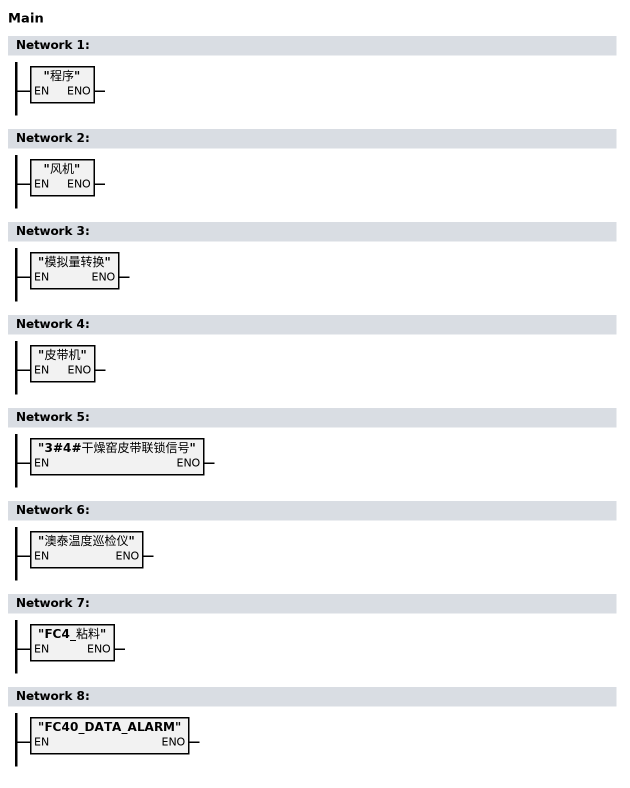
   RUNG wire#powerrail
      "程序"()
   END_RUNG
   // the same network as SCL:
   "程序"();
END_REGION

REGION Network 2
   RUNG wire#powerrail
      "风机"()
   END_RUNG
   // the same network as SCL:
   "风机"();
END_REGION

REGION Network 3
   RUNG wire#powerrail
      "模拟量转换"()
   END_RUNG
   // the same network as SCL:
   "模拟量转换"();
END_REGION

REGION Network 4
   RUNG wire#powerrail
      "皮带机"()
   END_RUNG
   // the same network as SCL:
   "皮带机"();
END_REGION

REGION Network 5
   RUNG wire#powerrail
      "3#4#干燥窑皮带联锁信号"()
   END_RUNG
   // the same network as SCL:
   "3#4#干燥窑皮带联锁信号"();
END_REGION

REGION Network 6
   RUNG wire#powerrail
      "澳泰温度巡检仪"()
   END_RUNG
   // the same network as SCL:
   "澳泰温度巡检仪"();
END_REGION

REGION Network 7
   RUNG wire#powerrail
      "FC4_粘料"()
   END_RUNG
   // the same network as SCL:
   "FC4_粘料"();
END_REGION

REGION Network 8
   RUNG wire#powerrail
      "FC40_DATA_ALARM"()
   END_RUNG
   // the same network as SCL:
   "FC40_DATA_ALARM"();
END_REGION
END_ORGANIZATION_BLOCK

ORGANIZATION_BLOCK "Cyclic interrupt"   // OB30, LAD, CyclicInterrupt
{ S7_Optimized_Access := 'TRUE' }
VERSION : 0.1
   VAR_INPUT
      Initial_Call : Bool;   // Initial call of this OB
      Event_Count : Int;   // Events discarded
   END_VAR
   VAR_TEMP   // added for the SCL form of the ladder/FBD networks
      _w1 : Bool;
      _w2 : Bool;
   END_VAR
BEGIN

REGION Network 1
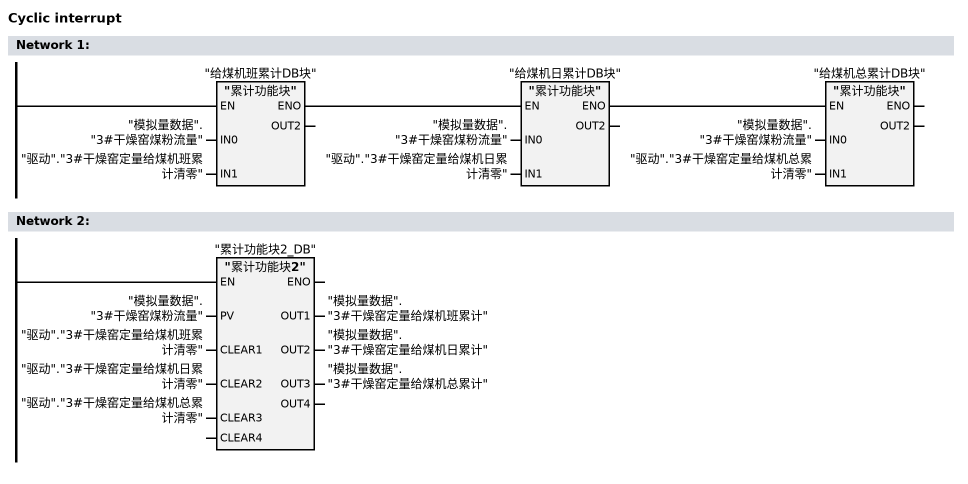
   RUNG wire#powerrail
      "给煤机班累计DB块"(IN0 := "模拟量数据"."3#干燥窑煤粉流量", IN1 := "驱动"."3#干燥窑定量给煤机班累计清零", OUT2 =>)
      "给煤机日累计DB块"(IN0 := "模拟量数据"."3#干燥窑煤粉流量", IN1 := "驱动"."3#干燥窑定量给煤机日累计清零", OUT2 =>)
      "给煤机总累计DB块"(IN0 := "模拟量数据"."3#干燥窑煤粉流量", IN1 := "驱动"."3#干燥窑定量给煤机总累计清零", OUT2 =>)
   END_RUNG
   // the same network as SCL:
   "给煤机班累计DB块"(IN0 := "模拟量数据"."3#干燥窑煤粉流量", IN1 := "驱动"."3#干燥窑定量给煤机班累计清零", ENO => #_w1);   // "累计功能块"
   "给煤机日累计DB块"(EN := #_w1, IN0 := "模拟量数据"."3#干燥窑煤粉流量", IN1 := "驱动"."3#干燥窑定量给煤机日累计清零", ENO => #_w2);   // "累计功能块"
   IF #_w2 THEN
       "给煤机总累计DB块"(IN0 := "模拟量数据"."3#干燥窑煤粉流量", IN1 := "驱动"."3#干燥窑定量给煤机总累计清零");   // "累计功能块"
   END_IF;
END_REGION

REGION Network 2
   RUNG wire#powerrail
      "累计功能块2_DB"(PV := "模拟量数据"."3#干燥窑煤粉流量", CLEAR1 := "驱动"."3#干燥窑定量给煤机班累计清零", CLEAR2 := "驱动"."3#干燥窑定量给煤机日累计清零", CLEAR3 := "驱动"."3#干燥窑定量给煤机总累计清零", CLEAR4 :=, OUT1 => "模拟量数据"."3#干燥窑定量给煤机班累计", OUT2 => "模拟量数据"."3#干燥窑定量给煤机日累计", OUT3 => "模拟量数据"."3#干燥窑定量给煤机总累计", OUT4 =>)
   END_RUNG
   // the same network as SCL:
   "累计功能块2_DB"(PV := "模拟量数据"."3#干燥窑煤粉流量",   // "累计功能块2"
               CLEAR1 := "驱动"."3#干燥窑定量给煤机班累计清零",
               CLEAR2 := "驱动"."3#干燥窑定量给煤机日累计清零",
               CLEAR3 := "驱动"."3#干燥窑定量给煤机总累计清零",
               OUT1 => "模拟量数据"."3#干燥窑定量给煤机班累计",
               OUT2 => "模拟量数据"."3#干燥窑定量给煤机日累计",
               OUT3 => "模拟量数据"."3#干燥窑定量给煤机总累计");
END_REGION
END_ORGANIZATION_BLOCK

// ===== PLC "3#HZY"  CPU 1511-1 PN =====

VAR_GLOBAL   // PLC tag table "默认变量表"
   "3#回转窑启动备妥" AT %I0.0 : Bool;
   "3#回转窑主机备妥" AT %I0.1 : Bool;
   "3#回转窑主机运行" AT %I0.2 : Bool;
   "3#回转窑主机故障" AT %I0.3 : Bool;
   "3#回转窑主机合闸" AT %I0.4 : Bool;
   "3#回转窑从机备妥" AT %I0.5 : Bool;
   "3#回转窑从机运行" AT %I0.6 : Bool;
   "3#回转窑从机故障" AT %I0.7 : Bool;
   "3#回转窑从机合闸" AT %I1.0 : Bool;
   "I1_3" AT %I1.3 : Bool;
   "I1_4" AT %I1.4 : Bool;
   "I1_5" AT %I1.5 : Bool;
   "I1_6" AT %I1.6 : Bool;
   "I1_7" AT %I1.7 : Bool;
   "主机稀油中控" AT %I2.0 : Bool;
   "主机稀油1#泵运行" AT %I2.1 : Bool;
   "主机稀油2#泵运行" AT %I2.2 : Bool;
   "主机稀油油差下限" AT %I2.3 : Bool;
   "主机稀油油位上限" AT %I2.4 : Bool;
   "主机稀油油位下限" AT %I2.5 : Bool;
   "主机稀油重故障" AT %I2.6 : Bool;
   "主机稀油轻故障" AT %I2.7 : Bool;
   "从机稀油中控" AT %I3.0 : Bool;
   "从机稀油1#泵运行" AT %I3.1 : Bool;
   "从机稀油2#泵运行" AT %I3.2 : Bool;
   "从机稀油油差下限" AT %I3.3 : Bool;
   "从机稀油油位上限" AT %I3.4 : Bool;
   "从机稀油油位下限" AT %I3.5 : Bool;
   "从机稀油重故障" AT %I3.6 : Bool;
   "从机稀油轻故障" AT %I3.7 : Bool;
   "1#挡轮备妥" AT %I4.0 : Bool;
   "1#挡轮1#泵运行" AT %I4.1 : Bool;
   "1#挡轮2#泵运行" AT %I4.2 : Bool;
   "1#挡轮溢流阀运行" AT %I4.3 : Bool;
   "挡轮重故障" AT %I4.4 : Bool;
   "挡轮轻故障" AT %I4.5 : Bool;
   "窑体行程上限" AT %I5.0 : Bool;
   "窑体行程上上限" AT %I5.1 : Bool;
   "窑体行程下限" AT %I5.2 : Bool;
   "窑体行程下下限" AT %I5.3 : Bool;
   "干矿提升皮带中控" AT %I6.0 : Bool;
   "干矿提升皮带运行" AT %I6.1 : Bool;
   "干矿提升皮带故障" AT %I6.2 : Bool;
   "干矿进料皮带中控" AT %I6.3 : Bool;
   "干矿进料皮带运行" AT %I6.4 : Bool;
   "干矿进料皮带故障" AT %I6.5 : Bool;
   "尾排风机高压远程" AT %I7.0 : Bool;
   "尾排风机高压合闸" AT %I7.1 : Bool;
   "尾排风机高压分闸" AT %I7.2 : Bool;
   "尾排风机变频远程" AT %I7.4 : Bool;
   "尾排风机变频运行" AT %I7.5 : Bool;
   "尾排风机变频故障" AT %I7.6 : Bool;
   "尾排风机变频待机" AT %I7.7 : Bool;
   "转子秤中控" AT %I8.0 : Bool;
   "转子秤运行" AT %I8.1 : Bool;
   "转子秤故障" AT %I8.2 : Bool;
   "煤粉仓收尘风机中控" AT %I8.4 : Bool;
   "煤粉仓收尘风机运行" AT %I8.5 : Bool;
   "煤粉仓收尘风机故障" AT %I8.6 : Bool;
   "回转窑一次风机中控" AT %I9.0 : Bool;
   "回转窑一次风机运行" AT %I9.1 : Bool;
   "回转窑一次风机故障" AT %I9.2 : Bool;
   "回转窑二次风机中控" AT %I9.3 : Bool;
   "回转窑二次风机运行" AT %I9.4 : Bool;
   "回转窑二次风机故障" AT %I9.5 : Bool;
   "回转窑备用一次风机中控" AT %I10.0 : Bool;
   "回转窑备用一次风机运行" AT %I10.1 : Bool;
   "回转窑备用一次风机故障" AT %I10.2 : Bool;
   "回转窑备用二次风机中控" AT %I10.3 : Bool;
   "回转窑备用二次风机运行" AT %I10.4 : Bool;
   "回转窑备用二次风机故障" AT %I10.5 : Bool;
   "回转窑窑头护板风机中控" AT %I11.0 : Bool;
   "回转窑窑头护板风机运行" AT %I11.1 : Bool;
   "回转窑窑头护板风机故障" AT %I11.2 : Bool;
   "回转窑助燃罗茨风机中控" AT %I11.3 : Bool;
   "回转窑助燃罗茨风机故障" AT %I11.4 : Bool;
   "回转窑助燃罗茨风机运行" AT %I11.5 : Bool;
   "23# 煤粉仓消防阀关到位" AT %I11.6 : Bool;
   "1#配料皮带备妥" AT %I12.0 : Bool;
   "1#配料皮带运行" AT %I12.1 : Bool;
   "1#配料皮带故障" AT %I12.2 : Bool;
   "1#配料皮带流量脉冲" AT %I12.3 : Bool;
   "2#配料皮带备妥" AT %I12.4 : Bool;
   "2#配料皮带运行" AT %I12.5 : Bool;
   "2#配料皮带故障" AT %I12.6 : Bool;
   "2#配料皮带流量脉冲" AT %I12.7 : Bool;
   "3#配料皮带备妥" AT %I13.0 : Bool;
   "3#配料皮带运行" AT %I13.1 : Bool;
   "3#配料皮带故障" AT %I13.2 : Bool;
   "3#配料皮带流量脉冲" AT %I13.3 : Bool;
   "4#配料皮带备妥" AT %I13.4 : Bool;
   "4#配料皮带运行" AT %I13.5 : Bool;
   "4#配料皮带故障" AT %I13.6 : Bool;
   "4#配料皮带流量脉冲" AT %I13.7 : Bool;
   "5#配料皮带备妥" AT %I14.0 : Bool;
   "5#配料皮带运行" AT %I14.1 : Bool;
   "5#配料皮带故障" AT %I14.2 : Bool;
   "5#配料皮带流量脉冲" AT %I14.3 : Bool;
   "6#配料皮带备妥" AT %I14.4 : Bool;
   "6#配料皮带运行" AT %I14.5 : Bool;
   "6#配料皮带故障" AT %I14.6 : Bool;
   "6#配料皮带流量脉冲" AT %I14.7 : Bool;
   "7#配料皮带备妥" AT %I15.0 : Bool;
   "7#配料皮带运行" AT %I15.1 : Bool;
   "7#配料皮带故障" AT %I15.2 : Bool;
   "7#配料皮带流量脉冲" AT %I15.3 : Bool;
   "1#板式给料机备妥" AT %I16.0 : Bool;
   "1#板式给料机运行" AT %I16.1 : Bool;
   "1#板式给料机故障" AT %I16.2 : Bool;
   "1#板式给料机流量脉冲" AT %I16.3 : Bool;
   "主机转速" AT %IW256 : Int;
   "主机电流" AT %IW258 : Int;
   "从机转速" AT %IW260 : Int;
   "从机电流" AT %IW262 : Int;
   "窑尾压力" AT %IW264 : Int;
   "尾排风机电流反馈" AT %IW266 : Int;
   "尾排风机频率反馈" AT %IW268 : Int;
   "烟道闸阀标尺" AT %IW270 : Int;
   "窑尾温度K偶" AT %IW280 : Int;
   "回转窑一次风机频率" AT %IW288 : Int;
   "回转窑一次风机电流" AT %IW290 : Int;
   "回转窑二次风机频率" AT %IW292 : Int;
   "回转窑二次风机电流" AT %IW294 : Int;
   "回转窑备用二次风机频率" AT %IW296 : Int;
   "回转窑备用二次风机电流" AT %IW298 : Int;
   "煤粉仓负压" AT %IW300 : Int;
   "转子秤流量反馈" AT %IW302 : Int;
   "回转窑窑头压力" AT %IW304 : Int;
   "一次风压力" AT %IW306 : Int;
   "二次风压力" AT %IW308 : Int;
   "煤粉仓温度1" AT %IW310 : Int;
   "煤粉仓温度2" AT %IW312 : Int;
   "煤粉仓温度3" AT %IW314 : Int;
   "煤粉仓温度4" AT %IW316 : Int;
   "回转窑助燃罗茨风机频率" AT %IW318 : Int;
   "回转窑助燃罗茨风机电流" AT %IW320 : Int;
   "窑头温度" AT %IW322 : Int;
   "窑体温度1" AT %IW324 : Int;
   "窑体温度2" AT %IW326 : Int;
   "窑体温度3" AT %IW328 : Int;
   "窑体温度4" AT %IW330 : Int;
   "窑体温度5" AT %IW332 : Int;
   "窑体温度6" AT %IW334 : Int;
   "1#配料流量" AT %IW336 : Int;
   "2#配料流量" AT %IW338 : Int;
   "3#配料流量" AT %IW340 : Int;
   "4#配料流量" AT %IW342 : Int;
   "3#回转窑支撑挡轮轴温度A1" AT %ID400 : DWord;
   "3#回转窑支撑挡轮温度A1" AT %ID404 : DWord;
   "3#回转窑支撑挡轮轴温度A2" AT %ID408 : DWord;
   "3#回转窑支撑挡轮温度A2" AT %ID412 : DWord;
   "3#回转窑支撑挡轮轴温度A3" AT %ID416 : DWord;
   "3#回转窑支撑挡轮温度A3" AT %ID420 : DWord;
   "3#回转窑支撑挡轮轴温度A4" AT %ID424 : DWord;
   "3#回转窑支撑挡轮温度A4" AT %ID428 : DWord;
   "3#回转窑支撑挡轮轴温度B1" AT %ID432 : DWord;
   "3#回转窑支撑挡轮温度B1" AT %ID436 : DWord;
   "3#回转窑支撑挡轮轴温度B2" AT %ID440 : DWord;
   "3#回转窑支撑挡轮温度B2" AT %ID444 : DWord;
   "3#回转窑支撑挡轮轴温度B3" AT %ID448 : DWord;
   "3#回转窑支撑挡轮温度B3" AT %ID452 : DWord;
   "3#回转窑支撑挡轮轴温度B4" AT %ID456 : DWord;
   "3#回转窑支撑挡轮温度B4" AT %ID460 : DWord;
   "3#回转窑支撑挡轮温度C1" AT %ID500 : DWord;
   "3#回转窑支撑挡轮轴温度C2" AT %ID504 : DWord;
   "3#回转窑支撑挡轮轴温度C3" AT %ID512 : DWord;
   "3#回转窑支撑挡轮温度C4" AT %ID524 : DWord;
   "3#回转窑支撑挡轮轴温度D1" AT %ID528 : DWord;
   "3#回转窑支撑挡轮温度D2" AT %ID540 : DWord;
   "3#回转窑支撑挡轮轴温度D3" AT %ID544 : DWord;
   "3#回转窑支撑挡轮轴温度D4" AT %ID552 : DWord;
   "3#回转窑支撑挡轮轴温度C1" AT %ID496 : DWord;
   "3#回转窑支撑挡轮温度C2" AT %ID508 : DWord;
   "3#回转窑支撑挡轮温度C3" AT %ID516 : DWord;
   "3#回转窑支撑挡轮轴温度C4" AT %ID520 : DWord;
   "3#回转窑支撑挡轮温度D1" AT %ID532 : DWord;
   "3#回转窑支撑挡轮轴温度D2" AT %ID536 : DWord;
   "3#回转窑支撑挡轮温度D3" AT %ID548 : DWord;
   "3#回转窑支撑挡轮温度D4" AT %ID556 : DWord;
   "3#回转窑煤粉仓称重" AT %ID600 : DWord;
   "3#回转窑中间仓称重" AT %ID608 : DWord;
   "转子秤流量脉冲" AT %I8.3 : Bool;
   "5#配料流量" AT %IW344 : Int;
   "6#配料流量" AT %IW346 : Int;
   "7#配料流量" AT %IW348 : Int;
   "板式给料机流量" AT %IW350 : Int;
   "3#窑提升皮带打滑信号" AT %I1.1 : Bool;
   "3#回转窑急停" AT %I1.2 : Bool;
   "I4_6" AT %I4.6 : Bool;
   "I4_7" AT %I4.7 : Bool;
   "主机稀油允许主机启动" AT %I5.4 : Bool;
   "从机稀油允许主机启动" AT %I5.5 : Bool;
   "I5_6" AT %I5.6 : Bool;
   "I5_7" AT %I5.7 : Bool;
   "I6_6" AT %I6.6 : Bool;
   "I6_7" AT %I6.7 : Bool;
   "I7_3" AT %I7.3 : Bool;
   "主电机定子温度" AT %IW272 : Int;
   "主电机前轴温度" AT %IW274 : Int;
   "主电机后轴温度" AT %IW276 : Int;
   "PIW278" AT %IW278 : Int;
   "从电机定子温度" AT %IW282 : Int;
   "从电机前轴温度" AT %IW284 : Int;
   "从电机后轴温度" AT %IW286 : Int;
   "I8_7" AT %I8.7 : Bool;
   "3#回转窑富氧快切阀开到位" AT %I9.6 : Bool;
   "3#回转窑富氧快切阀关到位" AT %I9.7 : Bool;
   "23# 煤粉仓消防阀自动位" AT %I10.6 : Bool;
   "23# 煤粉仓消防阀开到位" AT %I10.7 : Bool;
   "I11_7" AT %I11.7 : Bool;
   "I15_4" AT %I15.4 : Bool;
   "I15_5" AT %I15.5 : Bool;
   "I15_6" AT %I15.6 : Bool;
   "I15_7" AT %I15.7 : Bool;
   "I16_4" AT %I16.4 : Bool;
   "I16_5" AT %I16.5 : Bool;
   "I16_6" AT %I16.6 : Bool;
   "I16_7" AT %I16.7 : Bool;
   "I17_0" AT %I17.0 : Bool;
   "I17_1" AT %I17.1 : Bool;
   "I17_2" AT %I17.2 : Bool;
   "I17_3" AT %I17.3 : Bool;
   "I17_4" AT %I17.4 : Bool;
   "I17_5" AT %I17.5 : Bool;
   "I17_6" AT %I17.6 : Bool;
   "I17_7" AT %I17.7 : Bool;
   "回转窑合闸" AT %Q0.0 : Bool;
   "回转窑主机启动" AT %Q0.1 : Bool;
   "主机稀油启动" AT %Q0.2 : Bool;
   "从机稀油启动" AT %Q0.3 : Bool;
   "挡轮启动" AT %Q0.4 : Bool;
   "干矿提升皮带启动" AT %Q1.0 : Bool;
   "干矿进料皮带启动" AT %Q1.2 : Bool;
   "尾排风机高压合闸驱动" AT %Q1.3 : Bool;
   "尾排风机高压分闸驱动" AT %Q1.4 : Bool;
   "尾排风机高压柜变频启动" AT %Q1.5 : Bool;
   "尾排风机高压柜变频停止" AT %Q1.6 : Bool;
   "Q2_0" AT %Q2.0 : Bool;
   "Q2_1" AT %Q2.1 : Bool;
   "转子秤启动" AT %Q4.0 : Bool;
   "煤粉仓收尘风机启动" AT %Q4.1 : Bool;
   "回转窑一次风机启动" AT %Q4.2 : Bool;
   "回转窑二次风机启动" AT %Q4.3 : Bool;
   "回转窑备用一次风机启动" AT %Q4.4 : Bool;
   "回转窑备用二次风机启动" AT %Q4.5 : Bool;
   "回转窑窑头护板风机启动" AT %Q4.6 : Bool;
   "回转窑助燃罗茨风机启动" AT %Q4.7 : Bool;
   "转子秤连锁停止" AT %Q5.0 : Bool;
   "1#配料皮带启动" AT %Q6.0 : Bool;
   "2#配料皮带启动" AT %Q6.1 : Bool;
   "3#配料皮带启动" AT %Q6.2 : Bool;
   "4#配料皮带启动" AT %Q6.3 : Bool;
   "5#配料皮带启动" AT %Q6.4 : Bool;
   "6#配料皮带启动" AT %Q6.5 : Bool;
   "7#配料皮带启动" AT %Q6.6 : Bool;
   "板式给料机启动" AT %Q7.0 : Bool;
   "4#料仓粘仓信号输出" AT %Q7.1 : Bool;
   "Tag_34" AT %QB8 : Byte;
   "回转窑主机转速给定" AT %QW256 : Int;
   "尾排风机频率给定" AT %QW258 : Int;
   "给煤机流量给定" AT %QW272 : Int;
   "回转窑一次风机频率给定" AT %QW280 : Int;
   "回转窑二次风机频率给定" AT %QW282 : Int;
   "回转备用二次风机频率给定" AT %QW284 : Int;
   "1#配料流量给定" AT %QW288 : Int;
   "2#配料流量给定" AT %QW290 : Int;
   "3#配料流量给定" AT %QW292 : Int;
   "4#配料流量给定" AT %QW294 : Int;
   "5#配料流量给定" AT %QW296 : Int;
   "6#配料流量给定" AT %QW298 : Int;
   "7#配料流量给定" AT %QW300 : Int;
   "板式给料机流量给定" AT %QW302 : Int;
   "主机稀油停止" AT %Q0.5 : Bool;
   "从机稀油停止" AT %Q0.6 : Bool;
   "挡轮停止" AT %Q0.7 : Bool;
   "Q1_1" AT %Q1.1 : Bool;
   "Q1_7" AT %Q1.7 : Bool;
   "Q2_2" AT %Q2.2 : Bool;
   "Q2_3" AT %Q2.3 : Bool;
   "Q2_4" AT %Q2.4 : Bool;
   "Q2_5" AT %Q2.5 : Bool;
   "Q2_6" AT %Q2.6 : Bool;
   "Q2_7" AT %Q2.7 : Bool;
   "Q3_0" AT %Q3.0 : Bool;
   "Q3_1" AT %Q3.1 : Bool;
   "Q3_2" AT %Q3.2 : Bool;
   "Q3_3" AT %Q3.3 : Bool;
   "Q3_4" AT %Q3.4 : Bool;
   "Q3_5" AT %Q3.5 : Bool;
   "Q3_6" AT %Q3.6 : Bool;
   "Q3_7" AT %Q3.7 : Bool;
   "PQW260" AT %QW260 : Int;
   "PQW262" AT %QW262 : Int;
   "PQW264" AT %QW264 : Int;
   "PQW266" AT %QW266 : Int;
   "PQW268" AT %QW268 : Int;
   "PQW270" AT %QW270 : Int;
   "煤粉仓温度高报警" AT %Q5.1 : Bool;
   "23# 煤粉仓消防阀驱动" AT %Q5.2 : Bool;
   "Q5_3" AT %Q5.3 : Bool;
   "Q5_4" AT %Q5.4 : Bool;
   "Q5_5" AT %Q5.5 : Bool;
   "Q5_6" AT %Q5.6 : Bool;
   "3#回转窑富氧快切阀驱动" AT %Q5.7 : Bool;
   "3#回转窑富氧调节阀给定" AT %QW276 : Int;
   "PQW278" AT %QW278 : Int;
   "窑尾罩温度输出" AT %QW286 : Int;
   "Q6_7" AT %Q6.7 : Bool;
   "5#料仓粘仓信号输出" AT %Q7.2 : Bool;
   "6#料仓粘仓信号输出" AT %Q7.3 : Bool;
   "7#料仓粘仓信号输出" AT %Q7.4 : Bool;
   "1#料仓粘仓信号输出" AT %Q7.5 : Bool;
   "2#料仓粘仓信号输出" AT %Q7.6 : Bool;
   "3#料仓粘仓信号输出" AT %Q7.7 : Bool;
   "助燃罗茨风机频率给定" AT %QW274 : Int;
   "Tag_25" AT %M0.0 : Bool;
   "Tag_16" AT %M0.1 : Bool;
   "从机稀油油差下限停窑计时" AT %M0.3 : Bool;
   "主机稀油油位上限停窑计时" AT %M0.4 : Bool;
   "Tag_1" AT %MW4 : Word;
   "Tag_2" AT %MW6 : Word;
   "窑体行程上上限停窑计时" AT %M8.0 : Bool;
   "窑体行程下下限停窑计时" AT %M8.1 : Bool;
   "Tag_12" AT %MW60 : Word;
   "Tag_17" AT %MW62 : Word;
   "Tag_27" AT %MW68 : Word;
   "Tag_29" AT %MW72 : Word;
   "Tag_31" AT %MW74 : Word;
   "Tag_11" AT %M80.4 : Bool;
   "闸阀上限" AT %M80.6 : Bool;
   "闸阀下限" AT %M80.7 : Bool;
   "Tag_24" AT %MW100 : Word;
   "Tag_15" AT %M101.6 : Bool;
   "Tag_13" AT %M101.7 : Bool;
   "Tag_26" AT %MD328 : DWord;
   "Tag_28" AT %MD336 : DWord;
   "Tag_30" AT %MD338 : DWord;
   "Tag_19" AT %M400.0 : Bool;
   "Tag_23" AT %M400.2 : Bool;
   "Tag_21" AT %M400.5 : Bool;
   "Tag_22" AT %MW410 : Word;
   "Tag_35" AT %M99.0 : Bool;
   "Tag_37" AT %M88.0 : Bool;
   "主机稀油重故障_BOOL" AT %M10.0 : Bool;
   "从机稀油重故障_BOOL" AT %M10.1 : Bool;
   "挡轮油站重故障_BOOL" AT %M10.2 : Bool;
   "回转窑转子秤连锁" AT %M80.2 : Bool;
   "Tag_18" AT %M2.0 : Bool;
   "Tag_38" AT %M2.1 : Bool;
   "zhongjianzhi4_1" AT %MD420 : Real;
   "zhongjianzhi4_2" AT %MD424 : Real;
   "zhongjianzhi4_3" AT %MD428 : Real;
   "zhongjianzhi4_4" AT %MD432 : Real;
   "zhongjianzhi5_1" AT %MD436 : Real;
   "zhongjianzhi5_2" AT %MD440 : Real;
   "zhongjianzhi5_3" AT %MD444 : Real;
   "zhongjianzhi5_4" AT %MD448 : Real;
   "zhongjianzhi6_1" AT %MD452 : Real;
   "zhongjianzhi6_2" AT %MD456 : Real;
   "zhongjianzhi6_3" AT %MD460 : Real;
   "zhongjianzhi6_4" AT %MD464 : Real;
   "zhongjianzhi7_1" AT %MD468 : Real;
   "zhongjianzhi7_2" AT %MD472 : Real;
   "zhongjianzhi7_3" AT %MD476 : Real;
   "zhongjianzhi7_4" AT %MD480 : Real;
   "System_Byte" AT %MB1 : Byte;
   "FirstScan" AT %M1.0 : Bool;
   "DiagStatusUpdate" AT %M1.1 : Bool;
   "AlwaysTRUE" AT %M1.2 : Bool;
   "AlwaysFALSE" AT %M1.3 : Bool;
   "煤粉仓温度高报警中间量" AT %M102.0 : Bool;
   "煤粉仓温度高报警试验按钮" AT %M102.1 : Bool;
   "提升皮带打滑故障" AT %M9.0 : Bool;
   "提升皮带打滑故障复位" AT %M9.1 : Bool;
   "23# 煤粉仓消防阀开阀按钮" AT %M9.2 : Bool;
   "23# 煤粉仓消防阀关阀按钮" AT %M9.3 : Bool;
   "Tag_32" AT %T100 : Timer;
   "Tag_33" AT %T101 : Timer;
   "Tag_7" AT %T107 : Timer;
   "Tag_8" AT %T108 : Timer;
   "Tag_10" AT %T111 : Timer;
   "Tag_9" AT %T112 : Timer;
   "挡轮站启动时间" AT %T10 : Timer;
   "挡轮站停止时间" AT %T11 : Timer;
   "主稀油站启动时间" AT %T12 : Timer;
   "主稀油站停止时间" AT %T13 : Timer;
   "从稀油站启动时间" AT %T14 : Timer;
   "从稀油站停止时间" AT %T15 : Timer;
   "主机稀油重故障判断时间" AT %T20 : Timer;
   "从机稀油重故障判断时间" AT %T21 : Timer;
   "挡轮油站重故障判断时间" AT %T22 : Timer;
   "Tag_3" AT %T30 : Timer;
   "Tag_4" AT %T31 : Timer;
   "Tag_5" AT %T32 : Timer;
   "Tag_6" AT %T33 : Timer;
   "Tag_36" AT %T34 : Timer;
   "Tag_39" AT %T35 : Timer;
   "Tag_40" AT %T36 : Timer;
   "Tag_41" AT %T37 : Timer;
   "Tag_42" AT %T38 : Timer;
   "Tag_43" AT %T113 : Timer;
   "Tag_44" AT %T114 : Timer;
   "Tag_14" AT %C1 : Counter;
   "Tag_20" AT %C3 : Counter;
   "3#回转窑富氧压力" AT %IW354 : Int;
   "3#回转窑富氧流量" AT %IW356 : Int;
   "3#回转窑富氧流量调节阀反馈" AT %IW358 : Int;
   "3#回转窑富氧快切阀开按钮" AT %M9.4 : Bool;
   "3#回转窑富氧快切阀关按钮" AT %M9.5 : Bool;
   "3#回转窑富氧压力连锁点" AT %M9.6 : Bool;
   "3#回转窑富氧连锁投入与解除" AT %M9.7 : Bool;
   "Tag_45" AT %T115 : Timer;
END_VAR

DATA_BLOCK "DB块"   // DB1
{ S7_Optimized_Access := 'FALSE' }
VERSION : 0.1
   VAR
      STAT0 : Bool;
      STAT1 : Bool;
      STAT2 : Bool;
      STAT3_1 : Bool;
      STAT4_1 : Bool;
      STAT5_1 : Bool;
      "3#回转窑烟气管道闸板上限给定" : Real := 180.0;
      "3#回转窑烟气管道闸板下限给定" : Real := 5.0;
      定量给煤机班累计清零 : Bool;
      定量给煤机日累计清零 : Bool;
      定量给煤机总累计清零 : Bool;
   END_VAR
BEGIN
END_DATA_BLOCK

DATA_BLOCK "DB2_配料站清零按钮"   // DB2
{ S7_Optimized_Access := 'FALSE' }
VERSION : 0.1
   VAR
      "班01-1" : Bool;
      "班01-2" : Bool;
      "班01-3" : Bool;
      "班01-4" : Bool;
      "班01-5" : Bool;
      "班01-6" : Bool;
      "班01-7" : Bool;
      "班01-8" : Bool;
      "日01-1" : Bool;
      "日01-2" : Bool;
      "日01-3" : Bool;
      "日01-4" : Bool;
      "日01-5" : Bool;
      "日01-6" : Bool;
      "日01-7" : Bool;
      "日01-8" : Bool;
      "月01-1" : Bool;
      "月01-2" : Bool;
      "月01-3" : Bool;
      "月01-4" : Bool;
      "月01-5" : Bool;
      "月01-6" : Bool;
      "月01-7" : Bool;
      "月01-8" : Bool;
      "总01-1" : Bool;
      "总01-2" : Bool;
      "总01-3" : Bool;
      "总01-4" : Bool;
      "总01-5" : Bool;
      "总01-6" : Bool;
      "总01-7" : Bool;
      "总01-8" : Bool;
      备用1 : Bool;
      备用2 : Bool;
      备用3 : Bool;
      备用4 : Bool;
      备用5 : Bool;
      备用6 : Bool;
      备用7 : Bool;
      备用8 : Bool;
      备用9 : Bool;
      备用10 : Bool;
      备用11 : Bool;
      备用12 : Bool;
      备用13 : Bool;
      备用14 : Bool;
      备用15 : Bool;
      备用16 : Bool;
   END_VAR
BEGIN
END_DATA_BLOCK

DATA_BLOCK "给煤机班累计DB块"   // DB3
{ S7_Optimized_Access := 'FALSE' }
VERSION : 0.0
// stored: InstanceOfName 累计功能块
"累计功能块"
BEGIN
END_DATA_BLOCK

DATA_BLOCK "给煤机日累计DB块"   // DB4
{ S7_Optimized_Access := 'FALSE' }
VERSION : 0.0
// stored: InstanceOfName 累计功能块
"累计功能块"
BEGIN
END_DATA_BLOCK

DATA_BLOCK "给煤机总累计DB块"   // DB5
{ S7_Optimized_Access := 'FALSE' }
VERSION : 0.0
// stored: InstanceOfName 累计功能块
"累计功能块"
BEGIN
END_DATA_BLOCK

DATA_BLOCK "DB6_皮带秤粘料"   // DB6
{ S7_Optimized_Access := 'FALSE' }
VERSION : 0.1
   VAR
      转子秤给定反馈差值 : Real;
      转子秤给定反馈差值绝对值 : Real;
      real3 : Real;
      real4 : Real;
      real5 : Real;
      real6 : Real;
      real7 : Real;
      real8 : Real;
      real9 : Real;
      real10 : Real;
      real11 : Real;
      real12 : Real;
      real13 : Real;
      real14 : Real;
      real15 : Real;
      real16 : Real;
      real17 : Real;
      real18 : Real;
      real19 : Real;
      real20 : Real;
      转子秤粘料报警 : Bool;
      板式给料机粘料报警 : Bool;
      "1#配料皮带粘料报警" : Bool;
      "2#配料皮带粘料报警" : Bool;
      "3#配料皮带粘料报警" : Bool;
      "4#配料皮带粘料报警" : Bool;
      "5#配料皮带粘料报警" : Bool;
      "6#配料皮带粘料报警" : Bool;
      "7#配料皮带粘料报警" : Bool;
      bool10 : Bool;
      bool11 : Bool;
      bool12 : Bool;
      bool13 : Bool;
      bool14 : Bool;
      bool15 : Bool;
      bool16 : Bool;
      bool17 : Bool;
      bool18 : Bool;
      bool19 : Bool;
      bool20 : Bool;
      bool21 : Bool;
   END_VAR
BEGIN
END_DATA_BLOCK

DATA_BLOCK "DB10"   // DB10
{ S7_Optimized_Access := 'FALSE' }
VERSION : 0.1
   VAR
      "3#回转窑主传转速" : Real := 960.0;
      "3#回转窑主传电流" : Real := 101.7778;
      "3#回转窑主传转速给定" : Real := 960.0;
      STAT3 : Real;
      "3#回转窑从传转速" : Real := 960.0;
      "3#回转窑从传电流" : Real := 103.4074;
      STAT6 : Real;
      STAT7 : Real;
      "3#回转窑窑体温度1" : Real := 611.1111;
      "3#回转窑窑体温度2" : Real := 616.522;
      "3#回转窑窑体温度3" : Real := 494.2998;
      "3#回转窑窑体温度4" : Real := 357.7546;
      "3#回转窑窑体温度5" : Real := 226.9387;
      "3#回转窑窑体温度6" : Real;
      STAT14 : Real;
      STAT15 : Real;
      STAT16 : Real;
      STAT17 : Real;
      STAT18 : Real;
      STAT19 : Real;
      "3#回转窑窑尾温度" : Real := 307.3206;
      STAT21 : Real;
      "3#回转窑窑尾负压" : Real := -351.7361;
      STAT23 : Real;
      "3#回转窑煤粉仓温度1" : Real := 32.58102;
      "3#回转窑煤粉仓温度2" : Real := 32.58102;
      "3#回转窑煤粉仓温度3" : Real := 37.09491;
      "3#回转窑煤粉仓温度4" : Real := 33.73843;
      "3#回转窑煤粉仓温度5" : Real := 34.31713;
      "3#回转窑煤粉仓温度6" : Real := 67.27431;
      STAT30 : Real;
      STAT31 : Real;
      STAT32 : Real;
      "3#回转窑助燃罗茨风机运行频率" : Real;
      "3#回转窑助燃罗茨风机运行电流" : Real;
      "3#回转窑助燃罗茨风机频率给定" : Real;
      "3#回转窑转子秤流量" : Real := 3.821759;
      "3#回转窑转子秤流量给定" : Real := 1.0;
      "3#回转窑煤粉仓称重" : Real := 11.14;   // 3#回转窑煤粉仓称重
      STAT39 : Real;
      "3#回转窑送煤风机管道压力" : Real := 11.875;
      STAT41 : Real;
      "3#回转窑煤粉仓压力" : Real := -3259.896;
      STAT43 : Real;
      "3#回转窑窑头温度" : Real := 104.456;
      STAT45 : Real;
      "3#回转窑窑头负压" : Real := -168.2292;
      STAT47 : Real;
      "3#回转窑中间仓称重" : Real := 2.53;   // 3#回转窑中间仓称重
      STAT49 : Real;
      "3#回转窑送风风机管道压力" : Real := 12.70833;
      "3#回转窑一次风机频率给定" : Real := 40.0;
      "3#回转窑一次风机运行频率" : Real := 39.5544;
      "3#回转窑二次风机运行频率" : Real := 29.86111;
      "3#回转窑二次风机频率给定" : Real := 30.0;
      "3#回转窑备用二次风机运行频率" : Real := 0.1446759;
      "3#回转窑一次风机运行电流" : Real := 54.93055;
      "3#回转窑二次风机运行电流" : Real := 64.79948;
      "3#回转窑备用二次风机频率给定" : Real := 5.0;
      "3#回转窑备用二次风机运行电流" : Real := 0.3382523;
      "3#回转窑支撑挡轮温度A1" : Real := 36.0;
      "3#回转窑支撑挡轮温度A2" : Real := 35.0;
      "3#回转窑支撑挡轮温度A3" : Real := 35.0;
      "3#回转窑支撑挡轮温度A4" : Real := 34.0;
      "3#回转窑支撑挡轮温度B1" : Real := 33.0;
      "3#回转窑支撑挡轮温度B2" : Real := 36.0;
      "3#回转窑支撑挡轮温度B3" : Real := 38.0;
      "3#回转窑支撑挡轮温度B4" : Real := 35.0;
      "3#回转窑支撑挡轮温度C1" : Real := 36.0;
      "3#回转窑支撑挡轮温度C2" : Real := 34.0;
      "3#回转窑支撑挡轮温度C3" : Real := 39.0;
      "3#回转窑支撑挡轮温度C4" : Real := 37.0;
      "3#回转窑支撑挡轮温度D1" : Real := 36.0;
      "3#回转窑支撑挡轮温度D2" : Real := 33.0;
      "3#回转窑支撑挡轮温度D3" : Real := 42.0;
      "3#回转窑支撑挡轮温度D4" : Real := 34.0;
      "3#回转窑支撑挡轮轴温度A1" : Real := 35.0;
      "3#回转窑支撑挡轮轴温度A2" : Real := 39.0;
      "3#回转窑支撑挡轮轴温度A3" : Real := 35.0;
      "3#回转窑支撑挡轮轴温度A4" : Real := 34.0;
      "3#回转窑支撑挡轮轴温度B1" : Real := 33.0;
      "3#回转窑支撑挡轮轴温度B2" : Real := 16000.0;
      "3#回转窑支撑挡轮轴温度B3" : Real := 30.0;
      "3#回转窑支撑挡轮轴温度B4" : Real := 33.0;
      "3#回转窑支撑挡轮轴温度C1" : Real := 35.0;
      "3#回转窑支撑挡轮轴温度C2" : Real := 22.0;
      "3#回转窑支撑挡轮轴温度C3" : Real := 34.0;
      "3#回转窑支撑挡轮轴温度C4" : Real := 35.0;
      "3#回转窑支撑挡轮轴温度D1" : Real := 32.0;
      "3#回转窑支撑挡轮轴温度D2" : Real := 31.0;
      "3#回转窑支撑挡轮轴温度D3" : Real := 33.0;
      "3#回转窑支撑挡轮轴温度D4" : Real := 33.0;
      STAT92 : Real;
      STAT93 : Real;
      STAT94 : Real;
      STAT95 : Real;
      STAT96 : Real;
      STAT97 : Real;
      "3#回转窑窑尾烟气管道标尺高度" : Real := 75.4051;
      "3#回转窑定量给煤机班累计" : Real := 3039.521;
      "3#回转窑定量给煤机日累计" : Real := 3039.521;
      "3#回转窑定量给煤机总累计" : Real := 3039.521;
   END_VAR
BEGIN
END_DATA_BLOCK

DATA_BLOCK "DB12"   // DB12
{ S7_Optimized_Access := 'FALSE' }
VERSION : 0.1
   VAR
      "3#回转窑主传接触器合闸" : Bool;
      "3#回转窑主传接触器分闸" : Bool;
      "3#回转窑主传变频器启动" : Bool;
      "3#回转窑主传变频器停止" : Bool;
      "3#回转窑主机稀油站启动" : Bool;
      "3#回转窑主机稀油站停止" : Bool;
      "3#回转窑从机稀油站启动" : Bool;
      "3#回转窑从机稀油站停止" : Bool;
      STAT8 : Bool;
      STAT9 : Bool;
      STAT10 : Bool;
      STAT11 : Bool;
      STAT12 : Bool;
      STAT13 : Bool;
      STAT14 : Bool;
      STAT15 : Bool;
      "3#回转窑煤粉仓收尘风机启动" : Bool;
      "3#回转窑煤粉仓收尘风机停止" : Bool;
      "3#回转窑转子秤启动" : Bool;
      "3#回转窑转子秤停止" : Bool;
      STAT20 : Bool;
      STAT21 : Bool;
      STAT22 : Bool;
      STAT23 : Bool;
      "3#回转窑窑头护板风机启动" : Bool;
      "3#回转窑窑头护板风机停止" : Bool;
      STAT26 : Bool;
      STAT27 : Bool;
      STAT28 : Bool;
      STAT29 : Bool;
      STAT30 : Bool;
      STAT31 : Bool;
      STAT32 : Bool;
      STAT33 : Bool;
      "3#回转窑干矿提升皮带启动" : Bool;
      "3#回转窑干矿提升皮带停止" : Bool;
      STAT36 : Bool;
      STAT37 : Bool;
      "3#回转窑干矿进料皮带启动" : Bool;
      "3#回转窑干矿进料皮带停止" : Bool;
      STAT40 : Bool;
      STAT41 : Bool;
      STAT42 : Bool;
      STAT43 : Bool;
      STAT44 : Bool;
      STAT45 : Bool;
      "3#回转窑一次风机启动" : Bool;
      "3#回转窑一次风机停止" : Bool;
      "3#回转窑二次风机启动" : Bool;
      "3#回转窑二次风机停止" : Bool;
      "3#回转窑备用一次风机启动" : Bool;
      "3#回转窑备用一次风机停止" : Bool;
      "3#回转窑备用二次风机启动" : Bool;
      "3#回转窑备用二次风机停止" : Bool;
      STAT54 : Bool;
      STAT55 : Bool;
      "3#回转窑助燃罗茨风机启动" : Bool;
      "3#回转窑助燃罗茨风机停止" : Bool;
      STAT58 : Bool;
      STAT59 : Bool;
      "3#回转窑挡轮油站启动" : Bool;
      "3#回转窑挡轮油站停止" : Bool;
      STAT62 : Bool;
      STAT63 : Bool;
      "3#回转窑联锁解锁状态" : Bool := TRUE;
      STAT65 : Bool;
      "3#回转窑烟气管道闸板上升" : Bool;
      "3#回转窑烟气管道闸板下降" : Bool;
      STAT68 : Bool;
      STAT69 : Bool;
   END_VAR
BEGIN
END_DATA_BLOCK

DATA_BLOCK "DB20"   // DB20
{ S7_Optimized_Access := 'FALSE' }
VERSION : 0.1
   VAR
      STAT0 : Real := 0.004340278;
      STAT1 : Real := 1.762153;
      STAT2 : Real := 1.918403;
      STAT3 : Real := 41.19792;
      STAT4 : Real := 36.25;
      STAT5 : Real := 14.45313;
      STAT6 : Real := 0.02604167;
      STAT7 : Real;
      STAT8 : Real;
      STAT9 : Real;
      STAT10 : Real;
      STAT11 : Real;
      STAT12 : Real;
      STAT13 : Real;
      STAT14 : Real := 15.16204;
      STAT15 : Real;
      STAT16 : Real;
      STAT17 : Real := 1.8;
      STAT18 : Real := 1.9;
      STAT19 : Real := 42.75;
      STAT20 : Real := 38.0;
      STAT21 : Real := 14.25;
      STAT22 : Real;
      STAT23 : Real;
      STAT24 : Real;
      STAT25 : Real;
      STAT26 : Real;
      STAT27 : Real;
      STAT28 : Real;
      STAT29 : Real;
      STAT30 : Real := 100.0;
      STAT31 : Real;
      STAT32 : Real;
      STAT33 : Real;
      STAT34 : Real := 1111.676;
      STAT35 : Real := 1111.676;
      STAT36 : Real := 1.2;
      STAT37 : Real := 21.50005;
      STAT38 : Real := 1360.115;
      STAT39 : Real := 1360.115;
      STAT40 : Real := 1.2;
      STAT41 : Real := 22.70005;
      STAT42 : Real := 1629.349;
      STAT43 : Real := 1629.349;
      STAT44 : Real := 31.0;
      STAT45 : Real := 476.0;
      STAT46 : Real := 25807.0;
      STAT47 : Real := 25807.0;
      STAT48 : Real := 26.0;
      STAT49 : Real := 492.0;
      STAT50 : Real := 28773.0;
      STAT51 : Real := 28773.0;
      STAT52 : Real := 10.0;
      STAT53 : Real := 182.0;
      STAT54 : Real := 32564.0;
      STAT55 : Real := 32564.0;
      STAT56 : Real;
      STAT57 : Real;
      STAT58 : Real := 14053.0;
      STAT59 : Real := 14053.0;
      STAT60 : Real;
      STAT61 : Real;
      STAT62 : Real;
      STAT63 : Real;
      STAT64 : Real;
      STAT65 : Real;
      STAT66 : Real;
      STAT67 : Real;
      STAT68 : Real;
      STAT69 : Real;
      STAT70 : Real;
      STAT71 : Real;
      STAT72 : Real;
      STAT73 : Real;
      STAT74 : Real;
      STAT75 : Real;
      STAT76 : Real;
      STAT77 : Real;
      STAT78 : Real;
      STAT79 : Real;
      STAT80 : Real;
      STAT81 : Real;
      STAT82 : Real;
      STAT83 : Real;
      STAT84 : Real;
      STAT85 : Real;
      STAT86 : Real;
      STAT87 : Real;
      STAT88 : Real := 93.0;
      STAT89 : Real := 18593.0;
      STAT90 : Real := 18593.0;
      STAT91 : Real := 18593.0;
      STAT92 : Bool;
      STAT93 : Bool;
      STAT94 : Bool;
      STAT95 : Bool;
      STAT96 : Bool;
      STAT97 : Bool;
      STAT98 : Bool;
      STAT99 : Bool;
      STAT100 : Bool;
      STAT101 : Bool;
      STAT102 : Bool;
      STAT103 : Bool;
      STAT104 : Bool;
      STAT105 : Bool;
      STAT106 : Bool;
      STAT107 : Bool;
   END_VAR
BEGIN
END_DATA_BLOCK

DATA_BLOCK "DB22"   // DB22
{ S7_Optimized_Access := 'FALSE' }
VERSION : 0.1
   VAR
      STAT0 : Real := 43.92361;
      STAT1 : Real := 41.50752;
      STAT2 : Real := 41.0;
      STAT3 : Bool;
      STAT4 : Bool;
      STAT5 : Bool;
      STAT6 : Bool;
      STAT7 : Bool;
      STAT8 : Bool;
      STAT9 : Bool;
      STAT10 : Bool;
   END_VAR
BEGIN
END_DATA_BLOCK

DATA_BLOCK "数据块_电机温度"   // DB23
{ S7_Optimized_Access := 'FALSE' }
VERSION : 0.1
   VAR
      主机电机定子温度 : Real;
      主机电机前轴温度 : Real;
      主机电机后轴温度 : Real;
      从机电机定子温度 : Real;
      从机电机前轴温度 : Real;
      从机电机后轴温度 : Real;
      "3#回转窑富氧流量" : Real;
      "3#回转窑富氧调节阀反馈" : Real;
      "3#回转窑富氧调节阀给定" : Real;
      "3#回转窑富氧压力" : Real;
      "3#回转窑富氧压力设定" : Real;
   END_VAR
BEGIN
END_DATA_BLOCK

DATA_BLOCK "DB201"   // DB201
{ S7_Optimized_Access := 'FALSE' }
VERSION : 0.0
// stored: InstanceOfName 给料电机启动块
"给料电机启动块"
BEGIN
END_DATA_BLOCK

DATA_BLOCK "DB202"   // DB202
{ S7_Optimized_Access := 'FALSE' }
VERSION : 0.0
// stored: InstanceOfName 给料电机启动块
"给料电机启动块"
BEGIN
END_DATA_BLOCK

DATA_BLOCK "DB203"   // DB203
{ S7_Optimized_Access := 'FALSE' }
VERSION : 0.0
// stored: InstanceOfName 给料电机启动块
"给料电机启动块"
BEGIN
END_DATA_BLOCK

DATA_BLOCK "DB204"   // DB204
{ S7_Optimized_Access := 'FALSE' }
VERSION : 0.0
// stored: InstanceOfName 给料电机启动块
"给料电机启动块"
BEGIN
END_DATA_BLOCK

DATA_BLOCK "DB205"   // DB205
{ S7_Optimized_Access := 'FALSE' }
VERSION : 0.0
// stored: InstanceOfName 给料电机启动块
"给料电机启动块"
BEGIN
END_DATA_BLOCK

DATA_BLOCK "DB206"   // DB206
{ S7_Optimized_Access := 'FALSE' }
VERSION : 0.0
// stored: InstanceOfName 给料电机启动块
"给料电机启动块"
BEGIN
END_DATA_BLOCK

DATA_BLOCK "DB207"   // DB207
{ S7_Optimized_Access := 'FALSE' }
VERSION : 0.0
// stored: InstanceOfName 给料电机启动块
"给料电机启动块"
BEGIN
END_DATA_BLOCK

DATA_BLOCK "DB208"   // DB208
{ S7_Optimized_Access := 'FALSE' }
VERSION : 0.0
// stored: InstanceOfName 给料电机启动块
"给料电机启动块"
BEGIN
END_DATA_BLOCK

DATA_BLOCK "DB210"   // DB210
{ S7_Optimized_Access := 'FALSE' }
VERSION : 0.0
// stored: InstanceOfName FB11
"FB11"
BEGIN
END_DATA_BLOCK

DATA_BLOCK "DB211"   // DB211
{ S7_Optimized_Access := 'FALSE' }
VERSION : 0.0
// stored: InstanceOfName FB11
"FB11"
BEGIN
END_DATA_BLOCK

DATA_BLOCK "DB212"   // DB212
{ S7_Optimized_Access := 'FALSE' }
VERSION : 0.0
// stored: InstanceOfName FB11
"FB11"
BEGIN
END_DATA_BLOCK

DATA_BLOCK "DB213"   // DB213
{ S7_Optimized_Access := 'FALSE' }
VERSION : 0.1
// stored: InstanceOfName FB11
"FB11"
BEGIN
END_DATA_BLOCK

DATA_BLOCK "DB214"   // DB214
{ S7_Optimized_Access := 'FALSE' }
VERSION : 0.1
// stored: InstanceOfName FB11
"FB11"
BEGIN
END_DATA_BLOCK

DATA_BLOCK "DB215"   // DB215
{ S7_Optimized_Access := 'FALSE' }
VERSION : 0.1
// stored: InstanceOfName FB11
"FB11"
BEGIN
END_DATA_BLOCK

DATA_BLOCK "DB216"   // DB216
{ S7_Optimized_Access := 'FALSE' }
VERSION : 0.1
// stored: InstanceOfName FB11
"FB11"
BEGIN
END_DATA_BLOCK

DATA_BLOCK "DB217"   // DB217
{ S7_Optimized_Access := 'FALSE' }
VERSION : 0.0
// stored: InstanceOfName FB9
"FB9"
BEGIN
END_DATA_BLOCK

DATA_BLOCK "DB218"   // DB218
{ S7_Optimized_Access := 'FALSE' }
VERSION : 0.1
// stored: InstanceOfName FB9
"FB9"
BEGIN
END_DATA_BLOCK

DATA_BLOCK "DB219"   // DB219
{ S7_Optimized_Access := 'FALSE' }
VERSION : 0.1
// stored: InstanceOfName FB9
"FB9"
BEGIN
END_DATA_BLOCK

DATA_BLOCK "DB220"   // DB220
{ S7_Optimized_Access := 'FALSE' }
VERSION : 0.0
// stored: InstanceOfName FB11
"FB11"
BEGIN
END_DATA_BLOCK

DATA_BLOCK "DB221"   // DB221
{ S7_Optimized_Access := 'FALSE' }
VERSION : 0.0
// stored: InstanceOfName FB11
"FB11"
BEGIN
END_DATA_BLOCK

DATA_BLOCK "DB222"   // DB222
{ S7_Optimized_Access := 'FALSE' }
VERSION : 0.0
// stored: InstanceOfName FB11
"FB11"
BEGIN
END_DATA_BLOCK

DATA_BLOCK "DB223"   // DB223
{ S7_Optimized_Access := 'FALSE' }
VERSION : 0.1
// stored: InstanceOfName FB9
"FB9"
BEGIN
END_DATA_BLOCK

DATA_BLOCK "DB224"   // DB224
{ S7_Optimized_Access := 'FALSE' }
VERSION : 0.1
// stored: InstanceOfName FB9
"FB9"
BEGIN
END_DATA_BLOCK

FUNCTION_BLOCK "FB1"   // FB1, LAD
{ S7_Optimized_Access := 'FALSE' }
VERSION : 0.1
   VAR_INPUT
      IN0 : Real;   // IN0
      IN1 : Bool;   // IN1
   END_VAR
   VAR_OUTPUT
      OUT2 : Real;   // OUT2
   END_VAR
   VAR
      STAT3 : Real;   // STAT3
      STAT4 : Real;   // STAT4
      STAT5 : Real;   // STAT5
   END_VAR
BEGIN

REGION Network 1
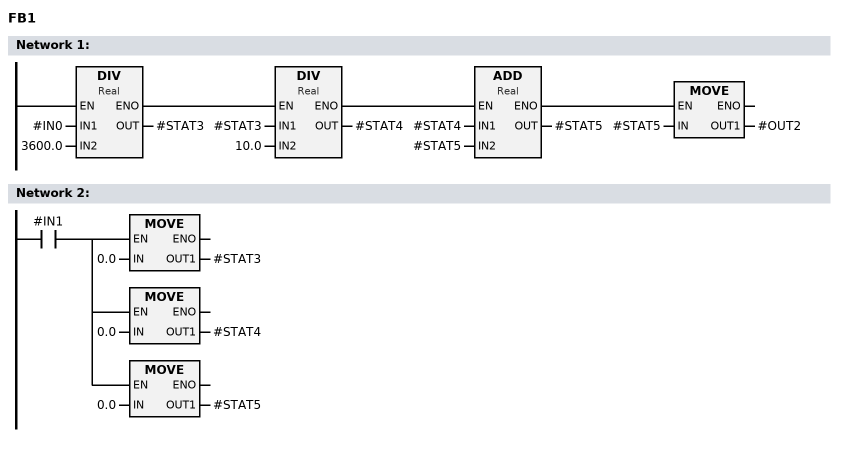
   RUNG wire#powerrail
      { S7_Templates := "SrcType := Real"; S7_GenerateENO := "TRUE" } Div(in1 := #IN0, in2 := 3600.0, out => #STAT3)
      { S7_Templates := "SrcType := Real"; S7_GenerateENO := "TRUE" } Div(in1 := #STAT3, in2 := 10.0, out => #STAT4)
      { S7_Templates := "SrcType := Real"; S7_GenerateENO := "TRUE" } Add(in1 := #STAT4, in2 := #STAT5, out => #STAT5)
      { S7_GenerateENO := "TRUE" } Move(in := #STAT5, out1 => #OUT2)
   END_RUNG
   // the same network as SCL:
   // ENO of a box is taken as its EN; it also drops when the box reports an error
   #STAT3 := #IN0 / 3600.0;
   #STAT4 := #STAT3 / 10.0;
   #STAT5 := #STAT4 + #STAT5;
   #OUT2 := #STAT5;
END_REGION

REGION Network 2
   RUNG wire#powerrail
      Contact( #IN1 )
      wire#w1
      { S7_GenerateENO := "TRUE" } Move(in := 0.0, out1 => #STAT3)
   END_RUNG
   RUNG wire#w1
      { S7_GenerateENO := "TRUE" } Move(in := 0.0, out1 => #STAT4)
   END_RUNG
   RUNG wire#w1
      { S7_GenerateENO := "TRUE" } Move(in := 0.0, out1 => #STAT5)
   END_RUNG
   // the same network as SCL:
   IF #IN1 THEN
       #STAT3 := 0.0;
       #STAT4 := 0.0;
       #STAT5 := 0.0;
   END_IF;
END_REGION
END_FUNCTION_BLOCK

FUNCTION_BLOCK "给料电机启动块"   // FB8, LAD
{ S7_Optimized_Access := 'FALSE' }
VERSION : 0.1
   VAR_INPUT
      IN0 : Bool;
      IN1 : Bool;
      IN2 : Bool;
      IN3 : Bool;
      IN4 : Bool;
      IN5 : Bool;
   END_VAR
   VAR_IN_OUT
      OUT6 : Bool;
   END_VAR
BEGIN

REGION Network 1
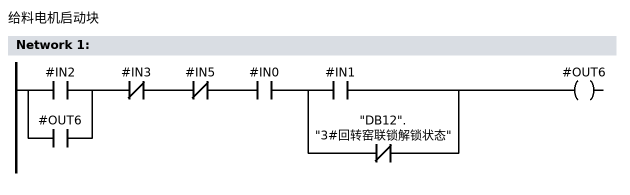
   RUNG wire#powerrail
      Contact( #IN2 )
      wire#w1
      I_Contact( #IN3 )
      I_Contact( #IN5 )
      Contact( #IN0 )
      wire#w2
      Contact( #IN1 )
      wire#w3
      Coil( #OUT6 )
   END_RUNG
   RUNG wire#powerrail
      Contact( #OUT6 )
   END_RUNG wire#w1
   RUNG wire#w2
      I_Contact( "DB12"."3#回转窑联锁解锁状态" )
   END_RUNG wire#w3
   // the same network as SCL:
   #OUT6 := (#IN2 OR #OUT6) AND NOT #IN3 AND NOT #IN5 AND #IN0 AND (#IN1 OR NOT "DB12"."3#回转窑联锁解锁状态");
END_REGION

REGION Network 2 (STL)
         SET;
         SAVE;
END_REGION
END_FUNCTION_BLOCK

FUNCTION_BLOCK "FB9"   // FB9, LAD
{ S7_Optimized_Access := 'FALSE' }